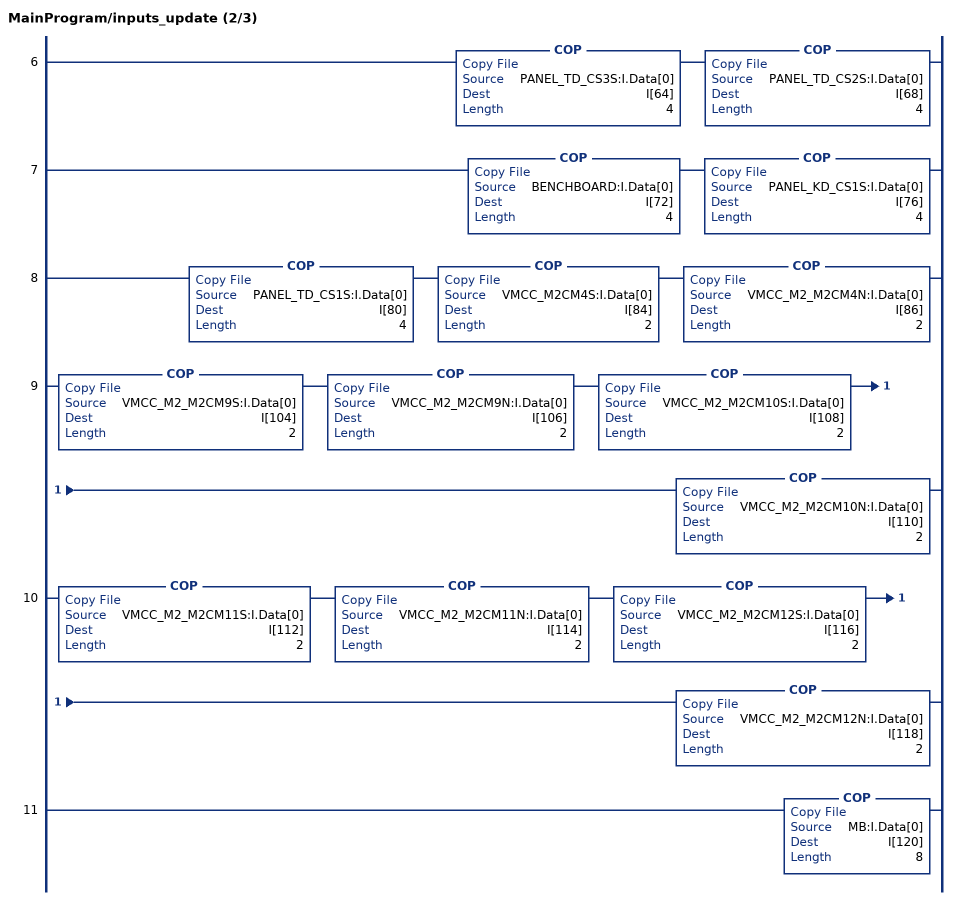
   6: COP(PANEL_TD_CS3S:I.Data[0],I[64],4)COP(PANEL_TD_CS2S:I.Data[0],I[68],4);
   7: COP(BENCHBOARD:I.Data[0],I[72],4)COP(PANEL_KD_CS1S:I.Data[0],I[76],4);
   8: COP(PANEL_TD_CS1S:I.Data[0],I[80],4)COP(VMCC_M2CM4S:I.Data[0],I[84],2)COP(VMCC_M2_M2CM4N:I.Data[0],I[86],2);
   9: COP(VMCC_M2_M2CM9S:I.Data[0],I[104],2)COP(VMCC_M2_M2CM9N:I.Data[0],I[106],2)COP(VMCC_M2_M2CM10S:I.Data[0],I[108],2)COP(VMCC_M2_M2CM10N:I.Data[0],I[110],2);
   10: COP(VMCC_M2_M2CM11S:I.Data[0],I[112],2)COP(VMCC_M2_M2CM11N:I.Data[0],I[114],2)COP(VMCC_M2_M2CM12S:I.Data[0],I[116],2)COP(VMCC_M2_M2CM12N:I.Data[0],I[118],2);
   11: COP(MB:I.Data[0],I[120],8);
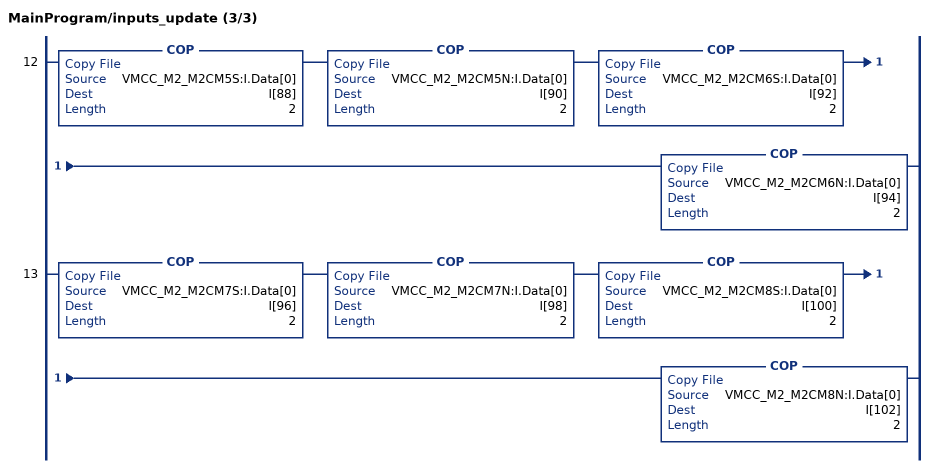
   12: COP(VMCC_M2_M2CM5S:I.Data[0],I[88],2)COP(VMCC_M2_M2CM5N:I.Data[0],I[90],2)COP(VMCC_M2_M2CM6S:I.Data[0],I[92],2)COP(VMCC_M2_M2CM6N:I.Data[0],I[94],2);
   13: COP(VMCC_M2_M2CM7S:I.Data[0],I[96],2)COP(VMCC_M2_M2CM7N:I.Data[0],I[98],2)COP(VMCC_M2_M2CM8S:I.Data[0],I[100],2)COP(VMCC_M2_M2CM8N:I.Data[0],I[102],2);
END_ROUTINE

ROUTINE M302SpeedUp_Faults   (* ladder *)
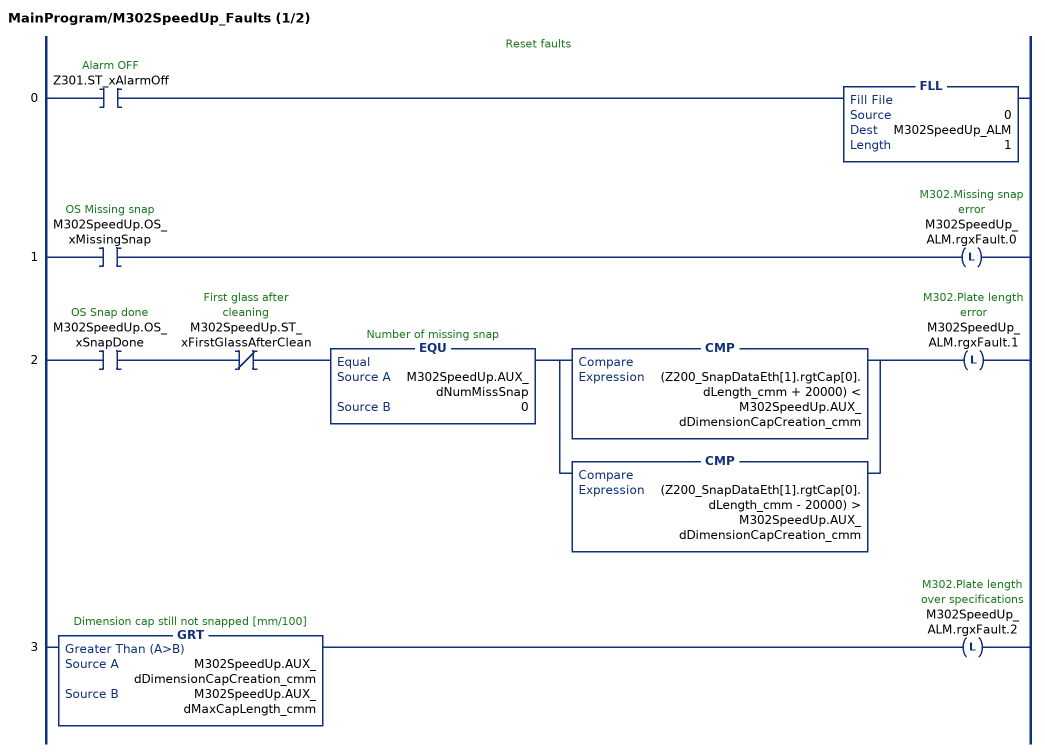
   // Reset faults
   0: XIC(Z301.ST_xAlarmOff)FLL(0,M302SpeedUp_ALM,1);
   1: XIC(M302SpeedUp.OS_xMissingSnap)OTL(M302SpeedUp_ALM.rgxFault.0);
   2: XIC(M302SpeedUp.OS_xSnapDone)XIO(M302SpeedUp.ST_xFirstGlassAfterClean)EQU(M302SpeedUp.AUX_dNumMissSnap,0)[CMP((Z200_SnapDataEth[1].rgtCap[0].dLength_cmm + 20000) < M302SpeedUp.AUX_dDimensionCapCreation_cmm) ,CMP((Z200_SnapDataEth[1].rgtCap[0].dLength_cmm - 20000) > M302SpeedUp.AUX_dDimensionCapCreation_cmm) ]OTL(M302SpeedUp_ALM.rgxFault.1);
   3: GRT(M302SpeedUp.AUX_dDimensionCapCreation_cmm,M302SpeedUp.AUX_dMaxCapLength_cmm)OTL(M302SpeedUp_ALM.rgxFault.2);
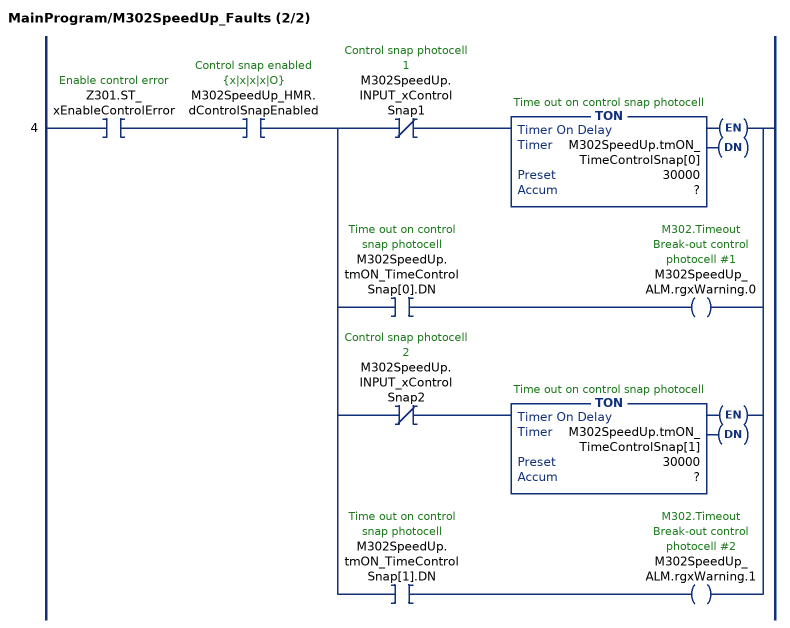
   4: XIC(Z301.ST_xEnableControlError)XIC(M302SpeedUp_HMR.dControlSnapEnabled)[XIO(M302SpeedUp.INPUT_xControlSnap1) TON(M302SpeedUp.tmON_TimeControlSnap[0],?,?) ,XIC(M302SpeedUp.tmON_TimeControlSnap[0].DN) OTE(M302SpeedUp_ALM.rgxWarning.0) ,XIO(M302SpeedUp.INPUT_xControlSnap2) TON(M302SpeedUp.tmON_TimeControlSnap[1],?,?) ,XIC(M302SpeedUp.tmON_TimeControlSnap[1].DN) OTE(M302SpeedUp_ALM.rgxWarning.1) ];
END_ROUTINE

ROUTINE M302SpeedUp_Logic   (* ladder *)
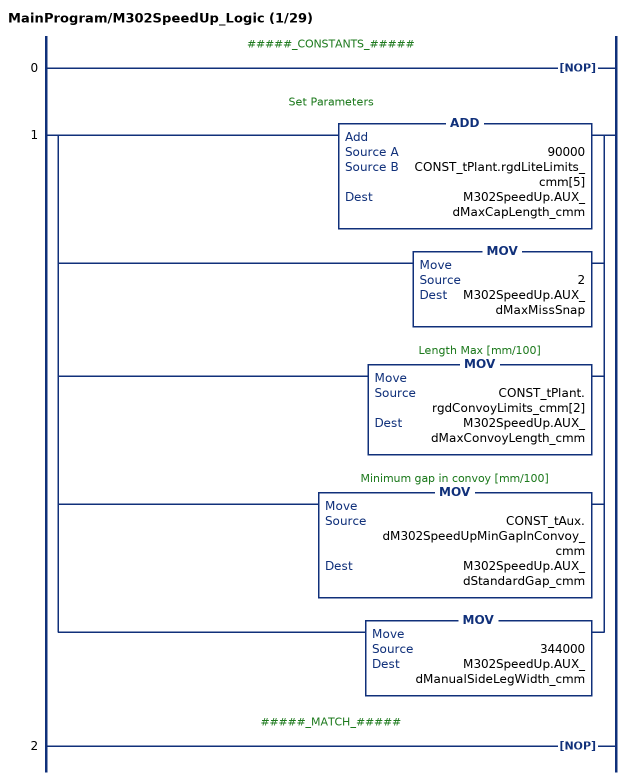
   // #####_CONSTANTS_#####
   0: NOP();
   // Set Parameters
   1: [ADD(90000,CONST_tPlant.rgdLiteLimits_cmm[5],M302SpeedUp.AUX_dMaxCapLength_cmm) ,MOV(2,M302SpeedUp.AUX_dMaxMissSnap) ,MOV(CONST_tPlant.rgdConvoyLimits_cmm[2],M302SpeedUp.AUX_dMaxConvoyLength_cmm) ,MOV(CONST_tAux.dM302SpeedUpMinGapInConvoy_cmm,M302SpeedUp.AUX_dStandardGap_cmm) ,MOV(344000,M302SpeedUp.AUX_dManualSideLegWidth_cmm) ];
   // #####_MATCH_#####
   2: NOP();
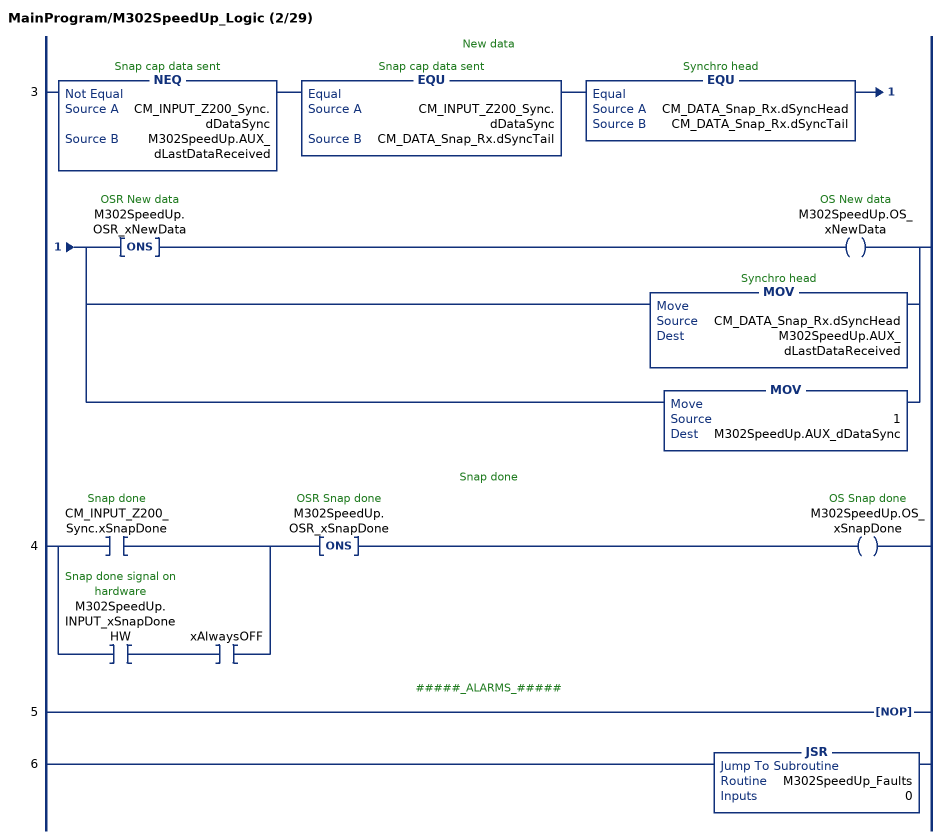
   // New data
   3: NEQ(CM_INPUT_Z200_Sync.dDataSync,M302SpeedUp.AUX_dLastDataReceived)EQU(CM_INPUT_Z200_Sync.dDataSync,CM_DATA_Snap_Rx.dSyncTail)EQU(CM_DATA_Snap_Rx.dSyncHead,CM_DATA_Snap_Rx.dSyncTail)[ONS(M302SpeedUp.OSR_xNewData) OTE(M302SpeedUp.OS_xNewData) ,MOV(CM_DATA_Snap_Rx.dSyncHead,M302SpeedUp.AUX_dLastDataReceived) ,MOV(1,M302SpeedUp.AUX_dDataSync) ];
   // Snap done
   4: [XIC(CM_INPUT_Z200_Sync.xSnapDone) ,XIC(M302SpeedUp.INPUT_xSnapDoneHW) XIC(xAlwaysOFF) ]ONS(M302SpeedUp.OSR_xSnapDone)OTE(M302SpeedUp.OS_xSnapDone);
   // #####_ALARMS_#####
   5: NOP();
   6: JSR(M302SpeedUp_Faults,0);
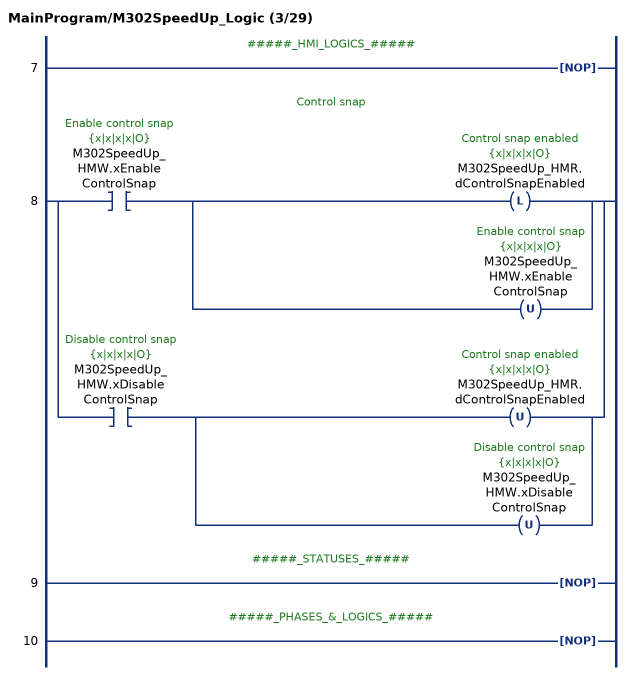
   // #####_HMI_LOGICS_#####
   7: NOP();
   // Control snap
   8: [XIC(M302SpeedUp_HMW.xEnableControlSnap) [OTL(M302SpeedUp_HMR.dControlSnapEnabled) ,OTU(M302SpeedUp_HMW.xEnableControlSnap) ] ,XIC(M302SpeedUp_HMW.xDisableControlSnap) [OTU(M302SpeedUp_HMR.dControlSnapEnabled) ,OTU(M302SpeedUp_HMW.xDisableControlSnap) ] ];
   // #####_STATUSES_#####
   9: NOP();
   // #####_PHASES_&_LOGICS_#####
   10: NOP();
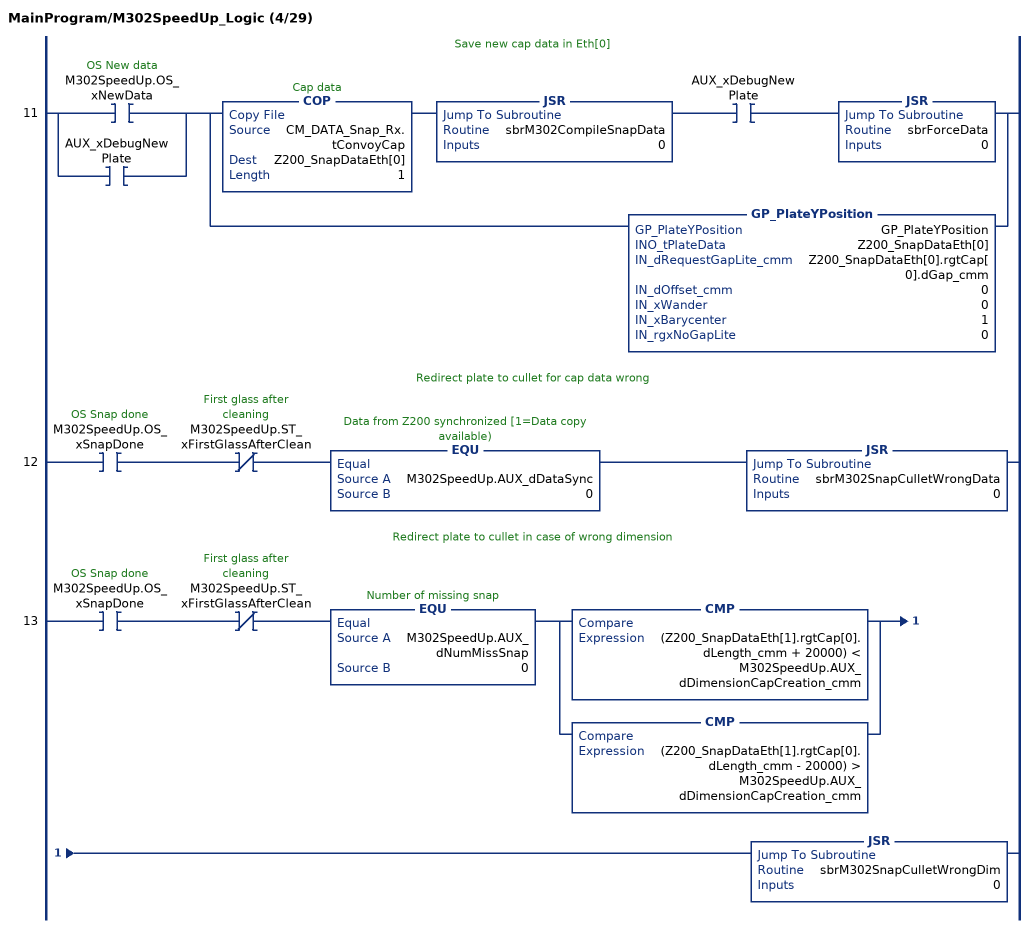
   // Save new cap data in Eth[0]
   11: [XIC(M302SpeedUp.OS_xNewData) ,XIC(AUX_xDebugNewPlate) ][COP(CM_DATA_Snap_Rx.tConvoyCap,Z200_SnapDataEth[0],1) JSR(sbrM302CompileSnapData,0) XIC(AUX_xDebugNewPlate) JSR(sbrForceData,0) ,GP_PlateYPosition(GP_PlateYPosition,Z200_SnapDataEth[0],Z200_SnapDataEth[0].rgtCap[0].dGap_cmm,0,0,1,0) ];
   // Redirect plate to cullet for cap data wrong
   12: XIC(M302SpeedUp.OS_xSnapDone)XIO(M302SpeedUp.ST_xFirstGlassAfterClean)EQU(M302SpeedUp.AUX_dDataSync,0)JSR(sbrM302SnapCulletWrongData,0);
   // Redirect plate to cullet in case of wrong dimension
   13: XIC(M302SpeedUp.OS_xSnapDone)XIO(M302SpeedUp.ST_xFirstGlassAfterClean)EQU(M302SpeedUp.AUX_dNumMissSnap,0)[CMP((Z200_SnapDataEth[1].rgtCap[0].dLength_cmm + 20000) < M302SpeedUp.AUX_dDimensionCapCreation_cmm) ,CMP((Z200_SnapDataEth[1].rgtCap[0].dLength_cmm - 20000) > M302SpeedUp.AUX_dDimensionCapCreation_cmm) ]JSR(sbrM302SnapCulletWrongDim,0);
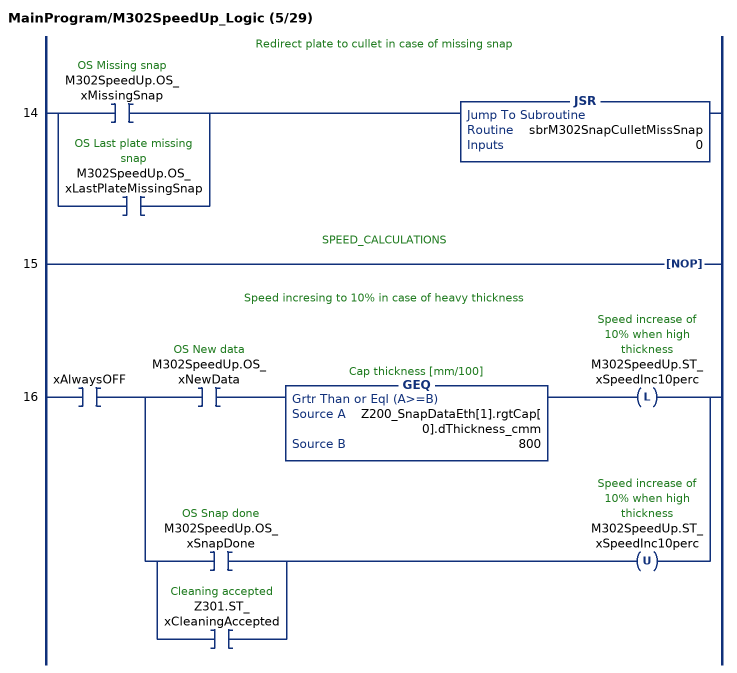
   // Redirect plate to cullet in case of missing snap
   14: [XIC(M302SpeedUp.OS_xMissingSnap) ,XIC(M302SpeedUp.OS_xLastPlateMissingSnap) ]JSR(sbrM302SnapCulletMissSnap,0);
   // SPEED_CALCULATIONS
   15: NOP();
   // Speed incresing to 10% in case of heavy thickness
   16: XIC(xAlwaysOFF)[XIC(M302SpeedUp.OS_xNewData) GEQ(Z200_SnapDataEth[1].rgtCap[0].dThickness_cmm,800) OTL(M302SpeedUp.ST_xSpeedInc10perc) ,[XIC(M302SpeedUp.OS_xSnapDone) ,XIC(Z301.ST_xCleaningAccepted) ] OTU(M302SpeedUp.ST_xSpeedInc10perc) ];
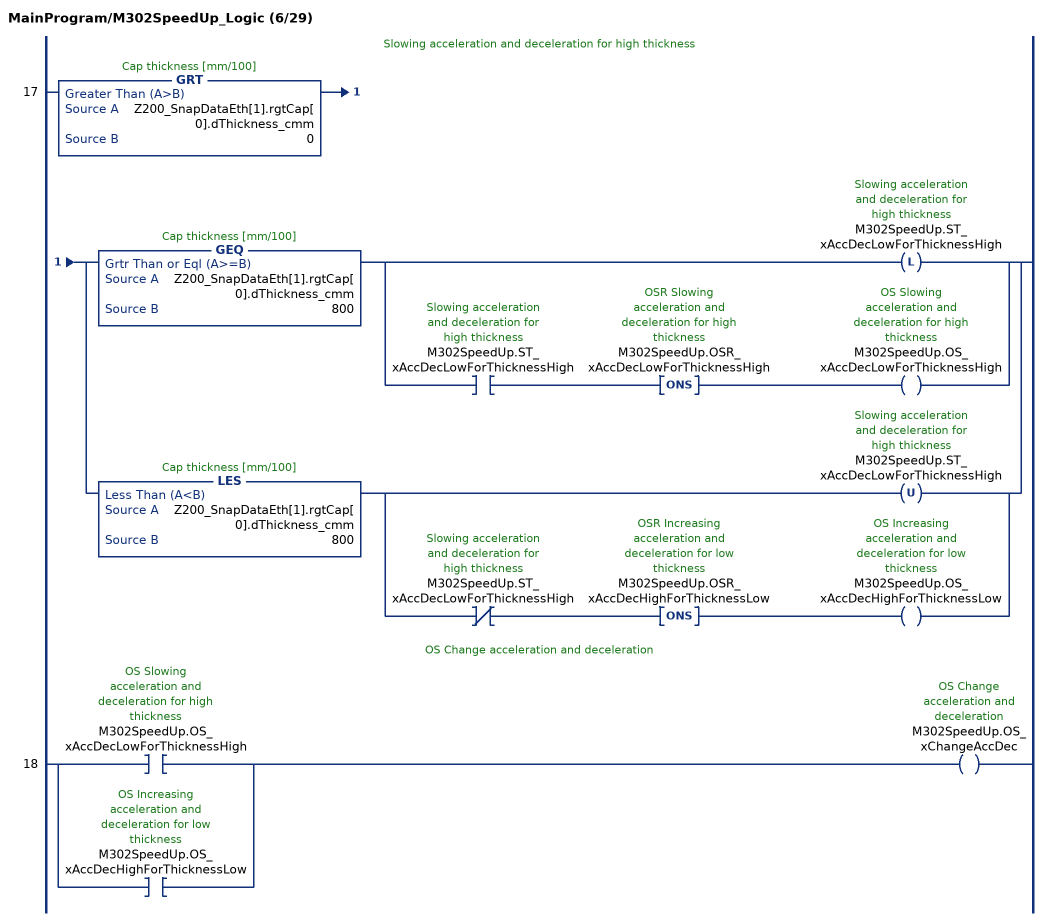
   // Slowing acceleration and deceleration for high thickness
   17: GRT(Z200_SnapDataEth[1].rgtCap[0].dThickness_cmm,0)[GEQ(Z200_SnapDataEth[1].rgtCap[0].dThickness_cmm,800) [OTL(M302SpeedUp.ST_xAccDecLowForThicknessHigh) ,XIC(M302SpeedUp.ST_xAccDecLowForThicknessHigh) ONS(M302SpeedUp.OSR_xAccDecLowForThicknessHigh) OTE(M302SpeedUp.OS_xAccDecLowForThicknessHigh) ] ,LES(Z200_SnapDataEth[1].rgtCap[0].dThickness_cmm,800) [OTU(M302SpeedUp.ST_xAccDecLowForThicknessHigh) ,XIO(M302SpeedUp.ST_xAccDecLowForThicknessHigh) ONS(M302SpeedUp.OSR_xAccDecHighForThicknessLow) OTE(M302SpeedUp.OS_xAccDecHighForThicknessLow) ] ];
   // OS Change acceleration and deceleration
   18: [XIC(M302SpeedUp.OS_xAccDecLowForThicknessHigh) ,XIC(M302SpeedUp.OS_xAccDecHighForThicknessLow) ]OTE(M302SpeedUp.OS_xChangeAccDec);
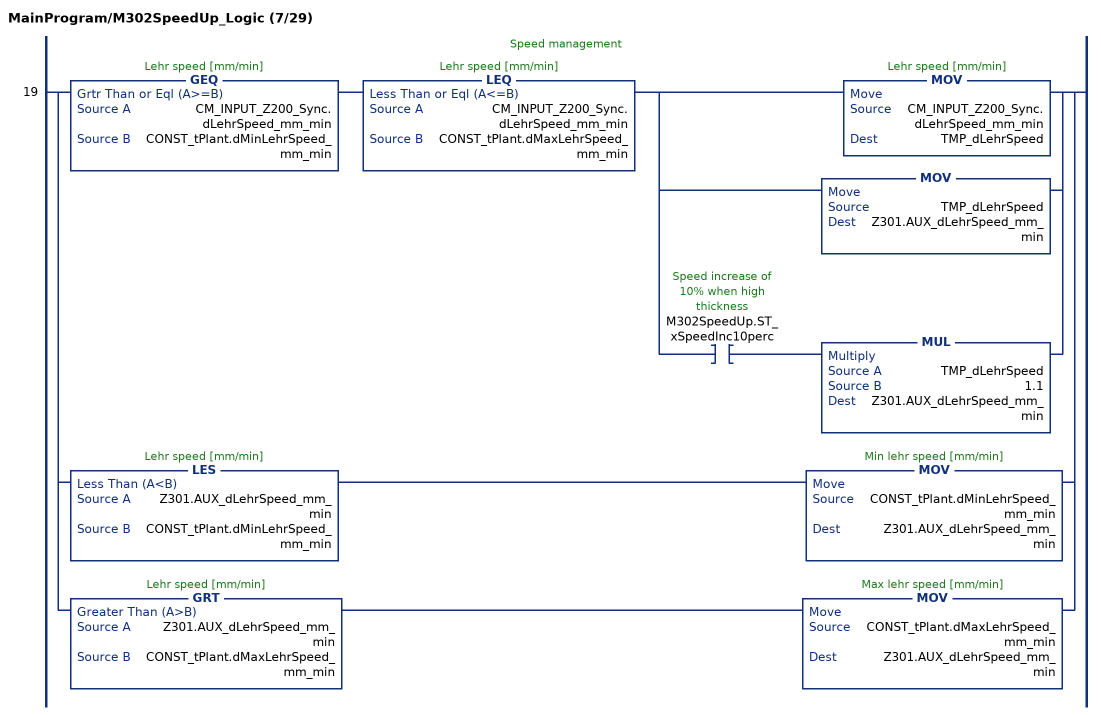
   // Speed management
   19: [GEQ(CM_INPUT_Z200_Sync.dLehrSpeed_mm_min,CONST_tPlant.dMinLehrSpeed_mm_min) LEQ(CM_INPUT_Z200_Sync.dLehrSpeed_mm_min,CONST_tPlant.dMaxLehrSpeed_mm_min) [MOV(CM_INPUT_Z200_Sync.dLehrSpeed_mm_min,TMP_dLehrSpeed) ,MOV(TMP_dLehrSpeed,Z301.AUX_dLehrSpeed_mm_min) ,XIC(M302SpeedUp.ST_xSpeedInc10perc) MUL(TMP_dLehrSpeed,1.1,Z301.AUX_dLehrSpeed_mm_min) ] ,LES(Z301.AUX_dLehrSpeed_mm_min,CONST_tPlant.dMinLehrSpeed_mm_min) MOV(CONST_tPlant.dMinLehrSpeed_mm_min,Z301.AUX_dLehrSpeed_mm_min) ,GRT(Z301.AUX_dLehrSpeed_mm_min,CONST_tPlant.dMaxLehrSpeed_mm_min) MOV(CONST_tPlant.dMaxLehrSpeed_mm_min,Z301.AUX_dLehrSpeed_mm_min) ];
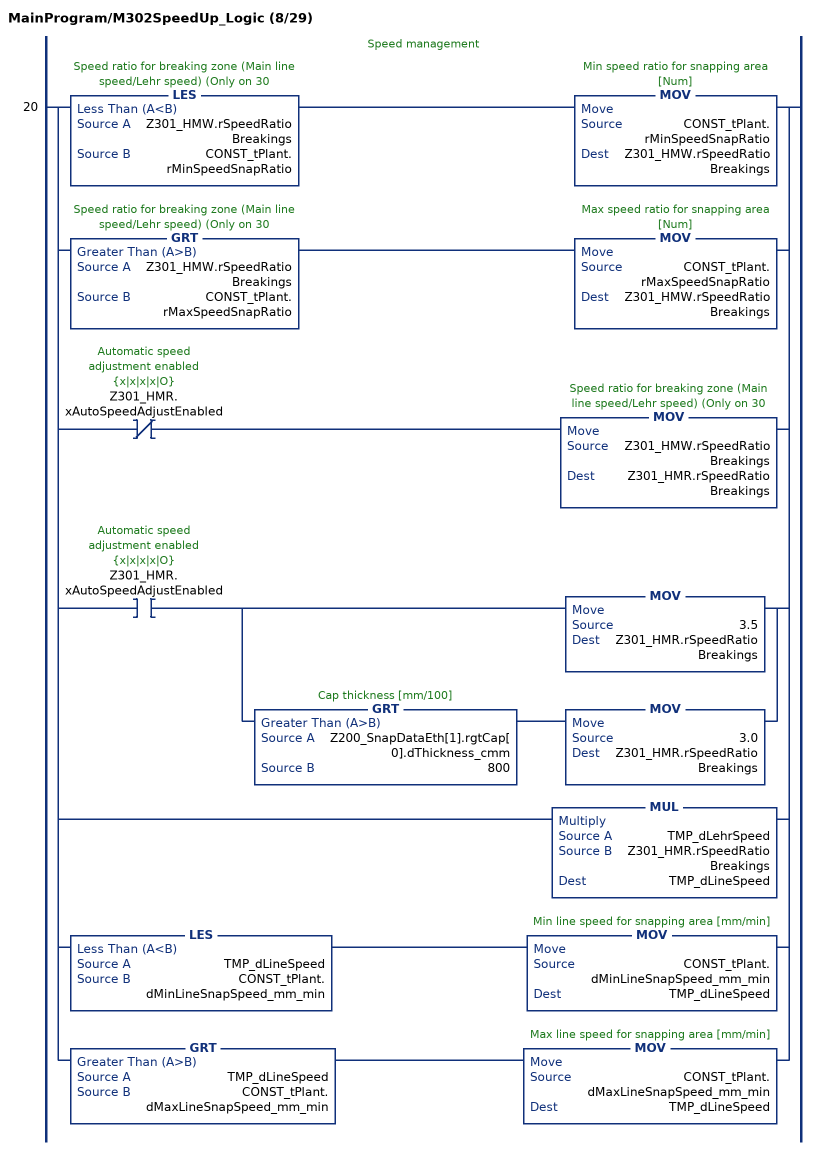
   // Speed management
   20: [LES(Z301_HMW.rSpeedRatioBreakings,CONST_tPlant.rMinSpeedSnapRatio) MOV(CONST_tPlant.rMinSpeedSnapRatio,Z301_HMW.rSpeedRatioBreakings) ,GRT(Z301_HMW.rSpeedRatioBreakings,CONST_tPlant.rMaxSpeedSnapRatio) MOV(CONST_tPlant.rMaxSpeedSnapRatio,Z301_HMW.rSpeedRatioBreakings) ,XIO(Z301_HMR.xAutoSpeedAdjustEnabled) MOV(Z301_HMW.rSpeedRatioBreakings,Z301_HMR.rSpeedRatioBreakings) ,XIC(Z301_HMR.xAutoSpeedAdjustEnabled) [MOV(3.5,Z301_HMR.rSpeedRatioBreakings) ,GRT(Z200_SnapDataEth[1].rgtCap[0].dThickness_cmm,800) MOV(3.0,Z301_HMR.rSpeedRatioBreakings) ] ,MUL(TMP_dLehrSpeed,Z301_HMR.rSpeedRatioBreakings,TMP_dLineSpeed) ,LES(TMP_dLineSpeed,CONST_tPlant.dMinLineSnapSpeed_mm_min) MOV(CONST_tPlant.dMinLineSnapSpeed_mm_min,TMP_dLineSpeed) ,GRT(TMP_dLineSpeed,CONST_tPlant.dMaxLineSnapSpeed_mm_min) MOV(CONST_tPlant.dMaxLineSnapSpeed_mm_min,TMP_dLineSpeed) ];
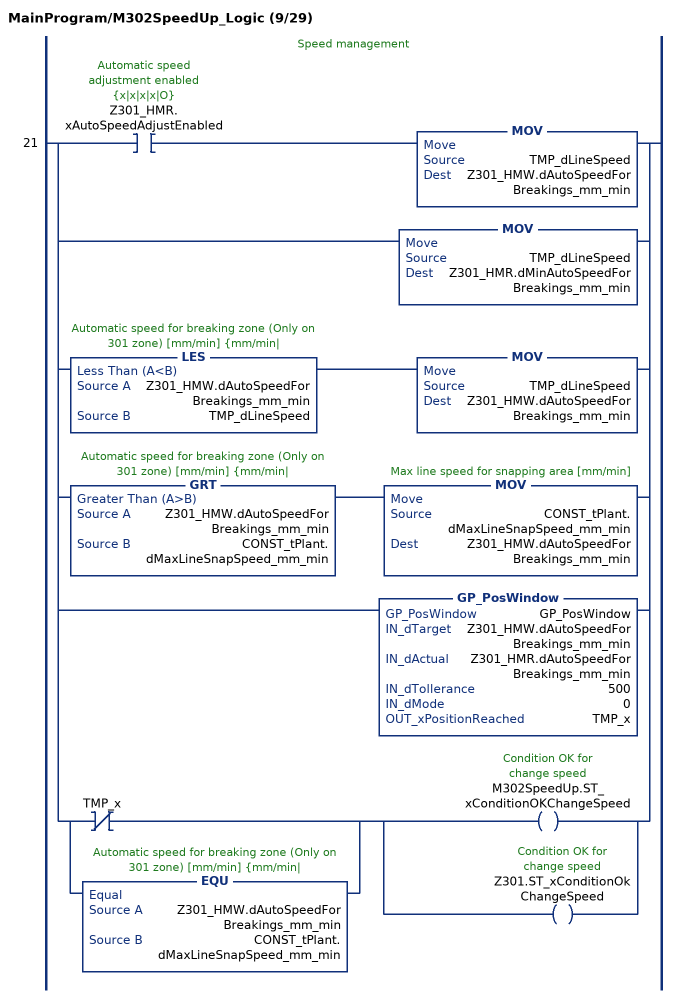
   // Speed management
   21: [XIC(Z301_HMR.xAutoSpeedAdjustEnabled) MOV(TMP_dLineSpeed,Z301_HMW.dAutoSpeedForBreakings_mm_min) ,MOV(TMP_dLineSpeed,Z301_HMR.dMinAutoSpeedForBreakings_mm_min) ,LES(Z301_HMW.dAutoSpeedForBreakings_mm_min,TMP_dLineSpeed) MOV(TMP_dLineSpeed,Z301_HMW.dAutoSpeedForBreakings_mm_min) ,GRT(Z301_HMW.dAutoSpeedForBreakings_mm_min,CONST_tPlant.dMaxLineSnapSpeed_mm_min) MOV(CONST_tPlant.dMaxLineSnapSpeed_mm_min,Z301_HMW.dAutoSpeedForBreakings_mm_min) ,[GP_PosWindow(GP_PosWindow,Z301_HMW.dAutoSpeedForBreakings_mm_min,Z301_HMR.dAutoSpeedForBreakings_mm_min,500,0,TMP_x) ,[XIO(TMP_x) ,EQU(Z301_HMW.dAutoSpeedForBreakings_mm_min,CONST_tPlant.dMaxLineSnapSpeed_mm_min) ] [OTE(M302SpeedUp.ST_xConditionOKChangeSpeed) ,OTE(Z301.ST_xConditionOkChangeSpeed) ] ] ];
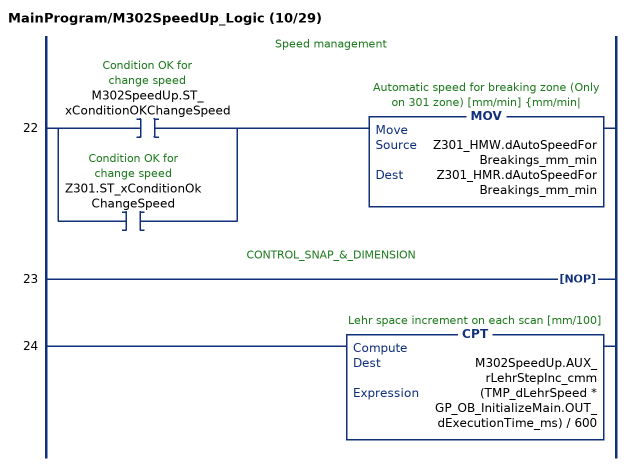
   // Speed management
   22: [XIC(M302SpeedUp.ST_xConditionOKChangeSpeed) ,XIC(Z301.ST_xConditionOkChangeSpeed) ]MOV(Z301_HMW.dAutoSpeedForBreakings_mm_min,Z301_HMR.dAutoSpeedForBreakings_mm_min);
   // CONTROL_SNAP_&_DIMENSION
   23: NOP();
   24: CPT(M302SpeedUp.AUX_rLehrStepInc_cmm,(TMP_dLehrSpeed * GP_OB_InitializeMain.OUT_dExecutionTime_ms) / 600);
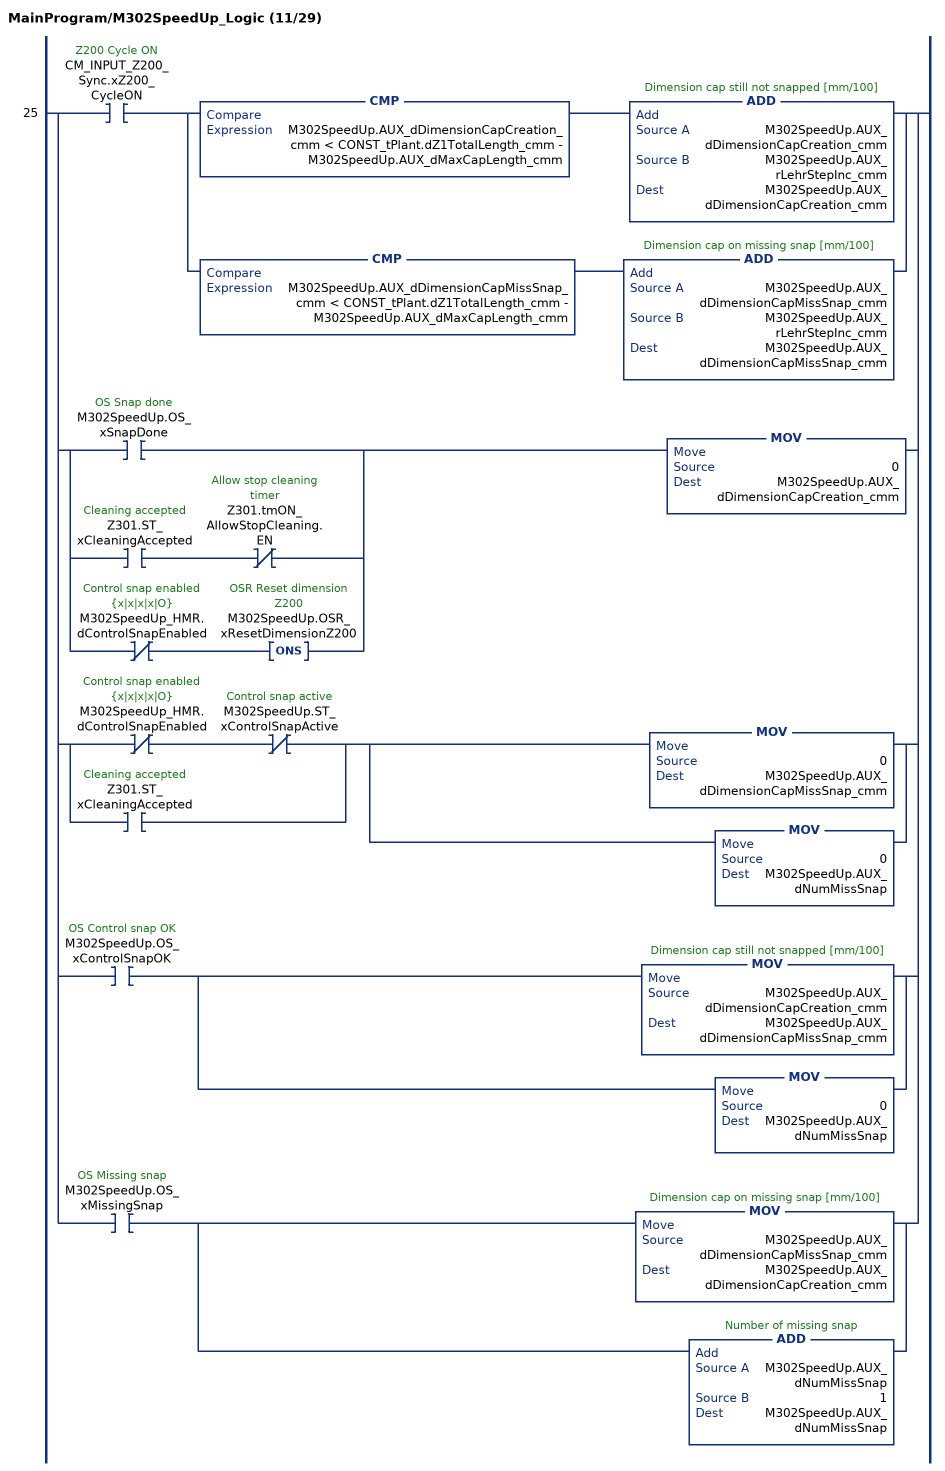
   25: [XIC(CM_INPUT_Z200_Sync.xZ200_CycleON) [CMP(M302SpeedUp.AUX_dDimensionCapCreation_cmm < CONST_tPlant.dZ1TotalLength_cmm - M302SpeedUp.AUX_dMaxCapLength_cmm) ADD(M302SpeedUp.AUX_dDimensionCapCreation_cmm,M302SpeedUp.AUX_rLehrStepInc_cmm,M302SpeedUp.AUX_dDimensionCapCreation_cmm) ,CMP(M302SpeedUp.AUX_dDimensionCapMissSnap_cmm < CONST_tPlant.dZ1TotalLength_cmm - M302SpeedUp.AUX_dMaxCapLength_cmm) ADD(M302SpeedUp.AUX_dDimensionCapMissSnap_cmm,M302SpeedUp.AUX_rLehrStepInc_cmm,M302SpeedUp.AUX_dDimensionCapMissSnap_cmm) ] ,[XIC(M302SpeedUp.OS_xSnapDone) ,XIC(Z301.ST_xCleaningAccepted) XIO(Z301.tmON_AllowStopCleaning.EN) ,XIO(M302SpeedUp_HMR.dControlSnapEnabled) ONS(M302SpeedUp.OSR_xResetDimensionZ200) ] MOV(0,M302SpeedUp.AUX_dDimensionCapCreation_cmm) ,[XIO(M302SpeedUp_HMR.dControlSnapEnabled) XIO(M302SpeedUp.ST_xControlSnapActive) ,XIC(Z301.ST_xCleaningAccepted) ] [MOV(0,M302SpeedUp.AUX_dDimensionCapMissSnap_cmm) ,MOV(0,M302SpeedUp.AUX_dNumMissSnap) ] ,XIC(M302SpeedUp.OS_xControlSnapOK) [MOV(M302SpeedUp.AUX_dDimensionCapCreation_cmm,M302SpeedUp.AUX_dDimensionCapMissSnap_cmm) ,MOV(0,M302SpeedUp.AUX_dNumMissSnap) ] ,XIC(M302SpeedUp.OS_xMissingSnap) [MOV(M302SpeedUp.AUX_dDimensionCapMissSnap_cmm,M302SpeedUp.AUX_dDimensionCapCreation_cmm) ,ADD(M302SpeedUp.AUX_dNumMissSnap,1,M302SpeedUp.AUX_dNumMissSnap) ] ];
